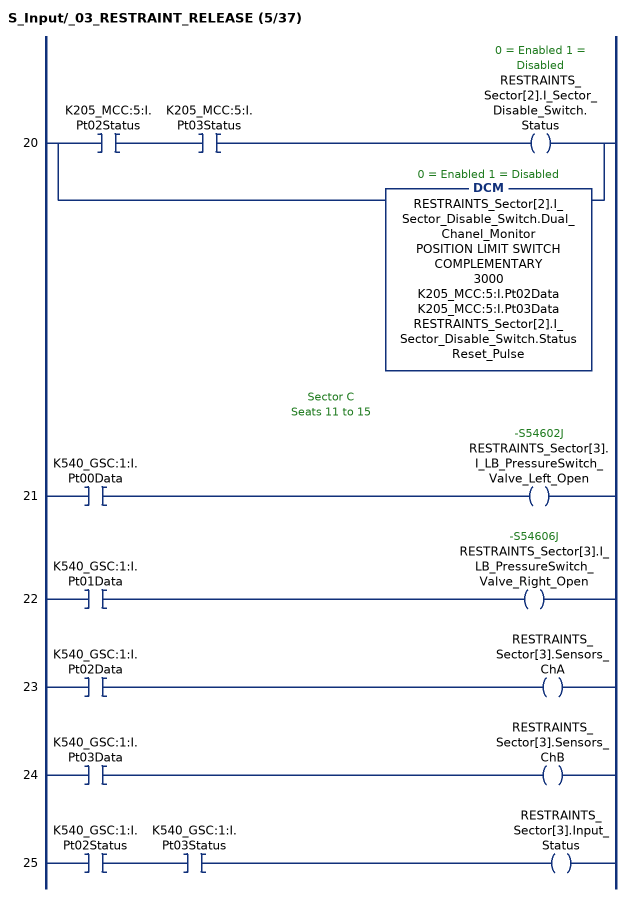
   20: [XIC(K205_MCC:5:I.Pt02Status) XIC(K205_MCC:5:I.Pt03Status) OTE(RESTRAINTS_Sector[2].I_Sector_Disable_Switch.Status) ,DCM(RESTRAINTS_Sector[2].I_Sector_Disable_Switch.Dual_Chanel_Monitor,POSITION LIMIT SWITCH,COMPLEMENTARY,3000,K205_MCC:5:I.Pt02Data,K205_MCC:5:I.Pt03Data,RESTRAINTS_Sector[2].I_Sector_Disable_Switch.Status,Reset_Pulse) ];
   // Sector C
   // Seats 11 to 15
   21: XIC(K540_GSC:1:I.Pt00Data)OTE(RESTRAINTS_Sector[3].I_LB_PressureSwitch_Valve_Left_Open);
   22: XIC(K540_GSC:1:I.Pt01Data)OTE(RESTRAINTS_Sector[3].I_LB_PressureSwitch_Valve_Right_Open);
   23: XIC(K540_GSC:1:I.Pt02Data)OTE(RESTRAINTS_Sector[3].Sensors_ChA);
   24: XIC(K540_GSC:1:I.Pt03Data)OTE(RESTRAINTS_Sector[3].Sensors_ChB);
   25: XIC(K540_GSC:1:I.Pt02Status)XIC(K540_GSC:1:I.Pt03Status)OTE(RESTRAINTS_Sector[3].Input_Status);
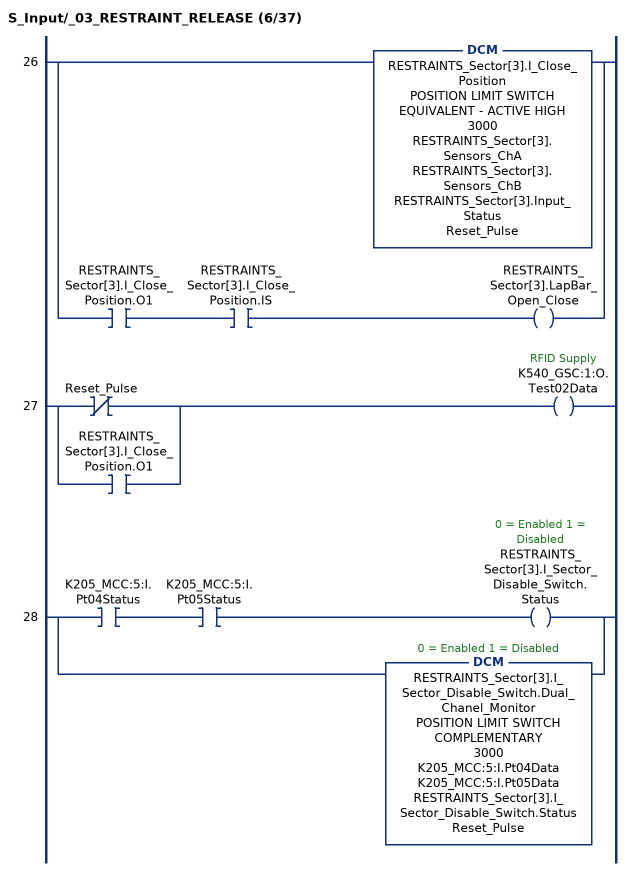
   26: [DCM(RESTRAINTS_Sector[3].I_Close_Position,POSITION LIMIT SWITCH,EQUIVALENT - ACTIVE HIGH,3000,RESTRAINTS_Sector[3].Sensors_ChA,RESTRAINTS_Sector[3].Sensors_ChB,RESTRAINTS_Sector[3].Input_Status,Reset_Pulse) ,XIC(RESTRAINTS_Sector[3].I_Close_Position.O1) XIC(RESTRAINTS_Sector[3].I_Close_Position.IS) OTE(RESTRAINTS_Sector[3].LapBar_Open_Close) ];
   27: [XIO(Reset_Pulse) ,XIC(RESTRAINTS_Sector[3].I_Close_Position.O1) ]OTE(K540_GSC:1:O.Test02Data);
   28: [XIC(K205_MCC:5:I.Pt04Status) XIC(K205_MCC:5:I.Pt05Status) OTE(RESTRAINTS_Sector[3].I_Sector_Disable_Switch.Status) ,DCM(RESTRAINTS_Sector[3].I_Sector_Disable_Switch.Dual_Chanel_Monitor,POSITION LIMIT SWITCH,COMPLEMENTARY,3000,K205_MCC:5:I.Pt04Data,K205_MCC:5:I.Pt05Data,RESTRAINTS_Sector[3].I_Sector_Disable_Switch.Status,Reset_Pulse) ];
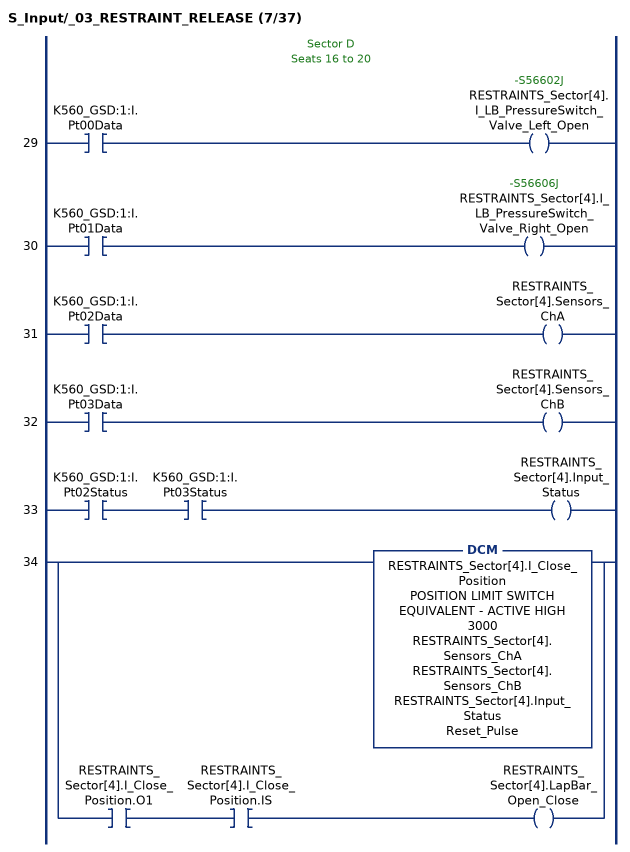
   // Sector D
   // Seats 16 to 20
   29: XIC(K560_GSD:1:I.Pt00Data)OTE(RESTRAINTS_Sector[4].I_LB_PressureSwitch_Valve_Left_Open);
   30: XIC(K560_GSD:1:I.Pt01Data)OTE(RESTRAINTS_Sector[4].I_LB_PressureSwitch_Valve_Right_Open);
   31: XIC(K560_GSD:1:I.Pt02Data)OTE(RESTRAINTS_Sector[4].Sensors_ChA);
   32: XIC(K560_GSD:1:I.Pt03Data)OTE(RESTRAINTS_Sector[4].Sensors_ChB);
   33: XIC(K560_GSD:1:I.Pt02Status)XIC(K560_GSD:1:I.Pt03Status)OTE(RESTRAINTS_Sector[4].Input_Status);
   34: [DCM(RESTRAINTS_Sector[4].I_Close_Position,POSITION LIMIT SWITCH,EQUIVALENT - ACTIVE HIGH,3000,RESTRAINTS_Sector[4].Sensors_ChA,RESTRAINTS_Sector[4].Sensors_ChB,RESTRAINTS_Sector[4].Input_Status,Reset_Pulse) ,XIC(RESTRAINTS_Sector[4].I_Close_Position.O1) XIC(RESTRAINTS_Sector[4].I_Close_Position.IS) OTE(RESTRAINTS_Sector[4].LapBar_Open_Close) ];
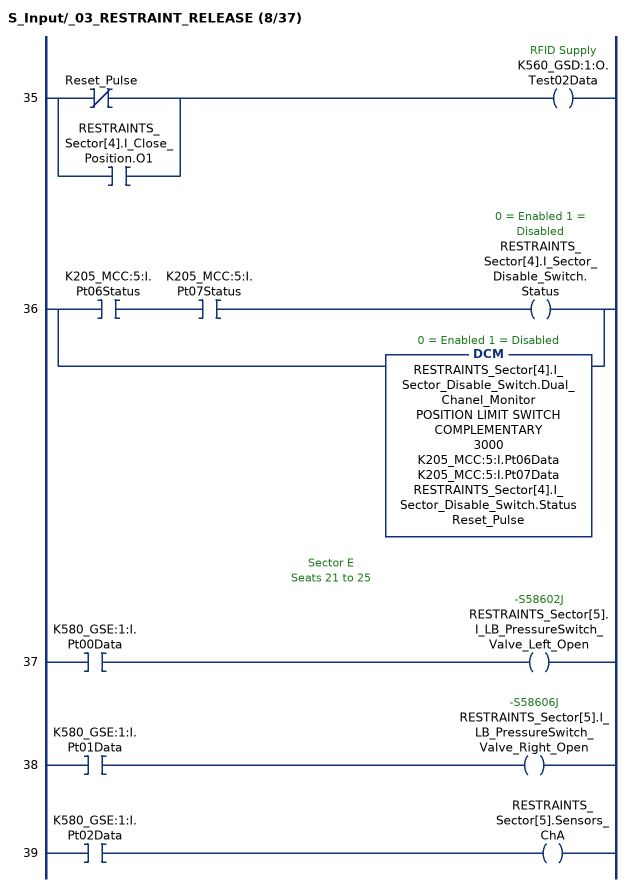
   35: [XIO(Reset_Pulse) ,XIC(RESTRAINTS_Sector[4].I_Close_Position.O1) ]OTE(K560_GSD:1:O.Test02Data);
   36: [XIC(K205_MCC:5:I.Pt06Status) XIC(K205_MCC:5:I.Pt07Status) OTE(RESTRAINTS_Sector[4].I_Sector_Disable_Switch.Status) ,DCM(RESTRAINTS_Sector[4].I_Sector_Disable_Switch.Dual_Chanel_Monitor,POSITION LIMIT SWITCH,COMPLEMENTARY,3000,K205_MCC:5:I.Pt06Data,K205_MCC:5:I.Pt07Data,RESTRAINTS_Sector[4].I_Sector_Disable_Switch.Status,Reset_Pulse) ];
   // Sector E
   // Seats 21 to 25
   37: XIC(K580_GSE:1:I.Pt00Data)OTE(RESTRAINTS_Sector[5].I_LB_PressureSwitch_Valve_Left_Open);
   38: XIC(K580_GSE:1:I.Pt01Data)OTE(RESTRAINTS_Sector[5].I_LB_PressureSwitch_Valve_Right_Open);
   39: XIC(K580_GSE:1:I.Pt02Data)OTE(RESTRAINTS_Sector[5].Sensors_ChA);
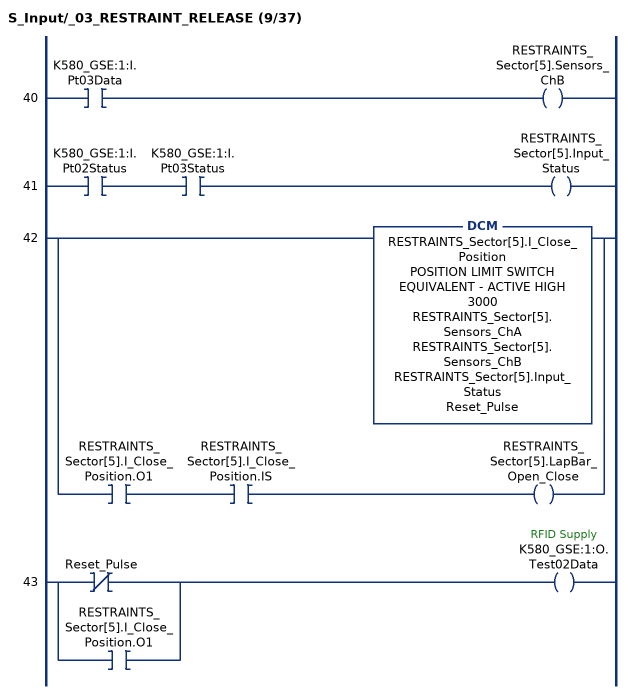
   40: XIC(K580_GSE:1:I.Pt03Data)OTE(RESTRAINTS_Sector[5].Sensors_ChB);
   41: XIC(K580_GSE:1:I.Pt02Status)XIC(K580_GSE:1:I.Pt03Status)OTE(RESTRAINTS_Sector[5].Input_Status);
   42: [DCM(RESTRAINTS_Sector[5].I_Close_Position,POSITION LIMIT SWITCH,EQUIVALENT - ACTIVE HIGH,3000,RESTRAINTS_Sector[5].Sensors_ChA,RESTRAINTS_Sector[5].Sensors_ChB,RESTRAINTS_Sector[5].Input_Status,Reset_Pulse) ,XIC(RESTRAINTS_Sector[5].I_Close_Position.O1) XIC(RESTRAINTS_Sector[5].I_Close_Position.IS) OTE(RESTRAINTS_Sector[5].LapBar_Open_Close) ];
   43: [XIO(Reset_Pulse) ,XIC(RESTRAINTS_Sector[5].I_Close_Position.O1) ]OTE(K580_GSE:1:O.Test02Data);
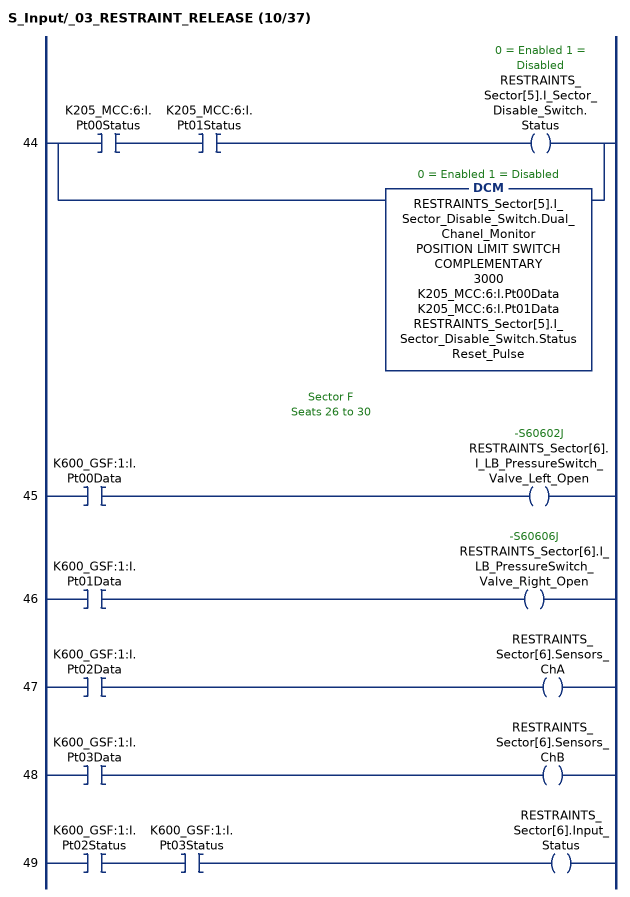
   44: [XIC(K205_MCC:6:I.Pt00Status) XIC(K205_MCC:6:I.Pt01Status) OTE(RESTRAINTS_Sector[5].I_Sector_Disable_Switch.Status) ,DCM(RESTRAINTS_Sector[5].I_Sector_Disable_Switch.Dual_Chanel_Monitor,POSITION LIMIT SWITCH,COMPLEMENTARY,3000,K205_MCC:6:I.Pt00Data,K205_MCC:6:I.Pt01Data,RESTRAINTS_Sector[5].I_Sector_Disable_Switch.Status,Reset_Pulse) ];
   // Sector F
   // Seats 26 to 30
   45: XIC(K600_GSF:1:I.Pt00Data)OTE(RESTRAINTS_Sector[6].I_LB_PressureSwitch_Valve_Left_Open);
   46: XIC(K600_GSF:1:I.Pt01Data)OTE(RESTRAINTS_Sector[6].I_LB_PressureSwitch_Valve_Right_Open);
   47: XIC(K600_GSF:1:I.Pt02Data)OTE(RESTRAINTS_Sector[6].Sensors_ChA);
   48: XIC(K600_GSF:1:I.Pt03Data)OTE(RESTRAINTS_Sector[6].Sensors_ChB);
   49: XIC(K600_GSF:1:I.Pt02Status)XIC(K600_GSF:1:I.Pt03Status)OTE(RESTRAINTS_Sector[6].Input_Status);
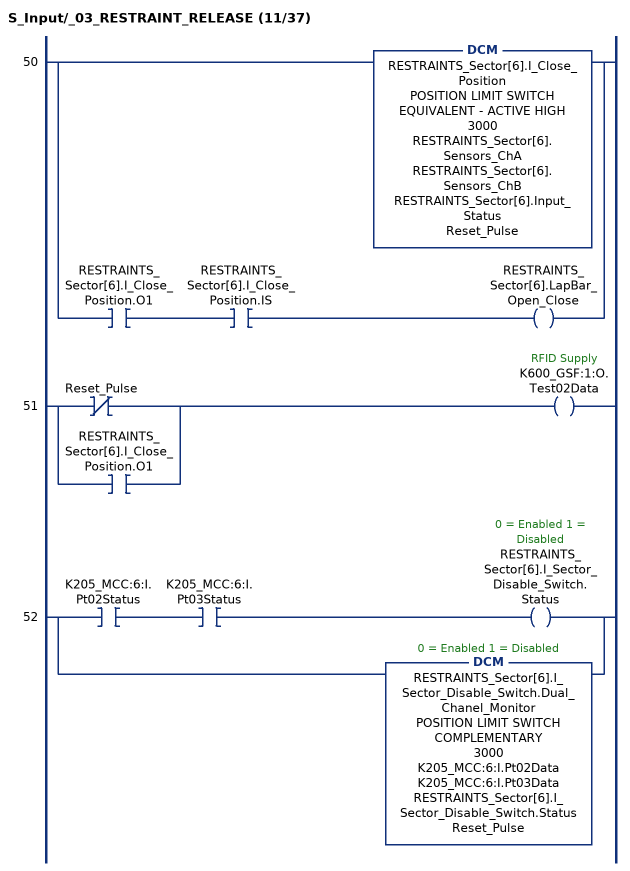
   50: [DCM(RESTRAINTS_Sector[6].I_Close_Position,POSITION LIMIT SWITCH,EQUIVALENT - ACTIVE HIGH,3000,RESTRAINTS_Sector[6].Sensors_ChA,RESTRAINTS_Sector[6].Sensors_ChB,RESTRAINTS_Sector[6].Input_Status,Reset_Pulse) ,XIC(RESTRAINTS_Sector[6].I_Close_Position.O1) XIC(RESTRAINTS_Sector[6].I_Close_Position.IS) OTE(RESTRAINTS_Sector[6].LapBar_Open_Close) ];
   51: [XIO(Reset_Pulse) ,XIC(RESTRAINTS_Sector[6].I_Close_Position.O1) ]OTE(K600_GSF:1:O.Test02Data);
   52: [XIC(K205_MCC:6:I.Pt02Status) XIC(K205_MCC:6:I.Pt03Status) OTE(RESTRAINTS_Sector[6].I_Sector_Disable_Switch.Status) ,DCM(RESTRAINTS_Sector[6].I_Sector_Disable_Switch.Dual_Chanel_Monitor,POSITION LIMIT SWITCH,COMPLEMENTARY,3000,K205_MCC:6:I.Pt02Data,K205_MCC:6:I.Pt03Data,RESTRAINTS_Sector[6].I_Sector_Disable_Switch.Status,Reset_Pulse) ];
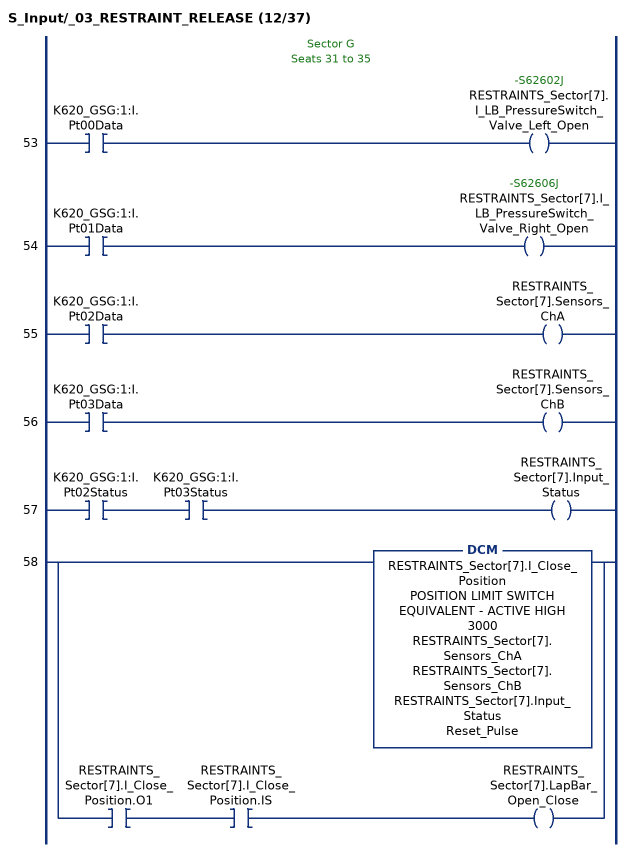
   // Sector G
   // Seats 31 to 35
   53: XIC(K620_GSG:1:I.Pt00Data)OTE(RESTRAINTS_Sector[7].I_LB_PressureSwitch_Valve_Left_Open);
   54: XIC(K620_GSG:1:I.Pt01Data)OTE(RESTRAINTS_Sector[7].I_LB_PressureSwitch_Valve_Right_Open);
   55: XIC(K620_GSG:1:I.Pt02Data)OTE(RESTRAINTS_Sector[7].Sensors_ChA);
   56: XIC(K620_GSG:1:I.Pt03Data)OTE(RESTRAINTS_Sector[7].Sensors_ChB);
   57: XIC(K620_GSG:1:I.Pt02Status)XIC(K620_GSG:1:I.Pt03Status)OTE(RESTRAINTS_Sector[7].Input_Status);
   58: [DCM(RESTRAINTS_Sector[7].I_Close_Position,POSITION LIMIT SWITCH,EQUIVALENT - ACTIVE HIGH,3000,RESTRAINTS_Sector[7].Sensors_ChA,RESTRAINTS_Sector[7].Sensors_ChB,RESTRAINTS_Sector[7].Input_Status,Reset_Pulse) ,XIC(RESTRAINTS_Sector[7].I_Close_Position.O1) XIC(RESTRAINTS_Sector[7].I_Close_Position.IS) OTE(RESTRAINTS_Sector[7].LapBar_Open_Close) ];
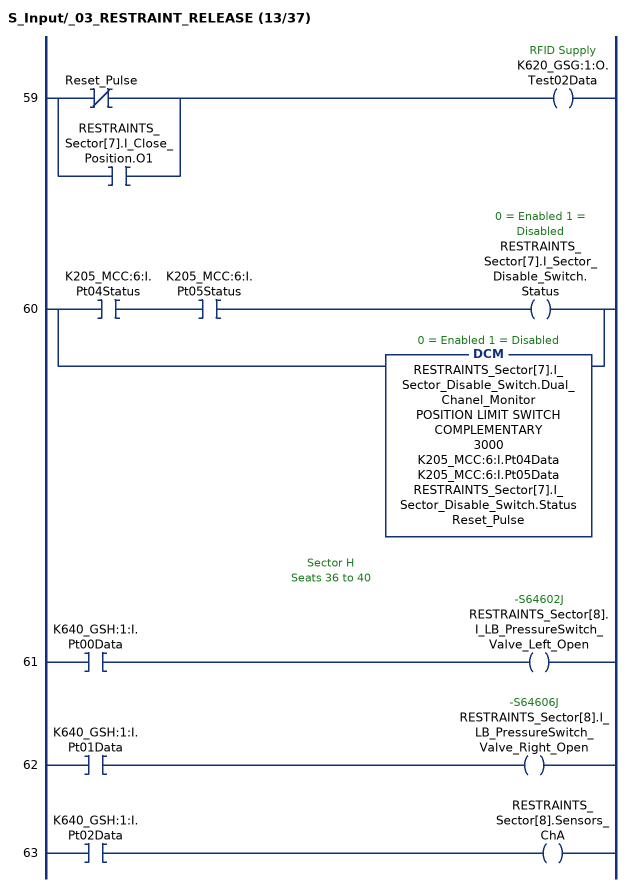
   59: [XIO(Reset_Pulse) ,XIC(RESTRAINTS_Sector[7].I_Close_Position.O1) ]OTE(K620_GSG:1:O.Test02Data);
   60: [XIC(K205_MCC:6:I.Pt04Status) XIC(K205_MCC:6:I.Pt05Status) OTE(RESTRAINTS_Sector[7].I_Sector_Disable_Switch.Status) ,DCM(RESTRAINTS_Sector[7].I_Sector_Disable_Switch.Dual_Chanel_Monitor,POSITION LIMIT SWITCH,COMPLEMENTARY,3000,K205_MCC:6:I.Pt04Data,K205_MCC:6:I.Pt05Data,RESTRAINTS_Sector[7].I_Sector_Disable_Switch.Status,Reset_Pulse) ];
   // Sector H
   // Seats 36 to 40
   61: XIC(K640_GSH:1:I.Pt00Data)OTE(RESTRAINTS_Sector[8].I_LB_PressureSwitch_Valve_Left_Open);
   62: XIC(K640_GSH:1:I.Pt01Data)OTE(RESTRAINTS_Sector[8].I_LB_PressureSwitch_Valve_Right_Open);
   63: XIC(K640_GSH:1:I.Pt02Data)OTE(RESTRAINTS_Sector[8].Sensors_ChA);
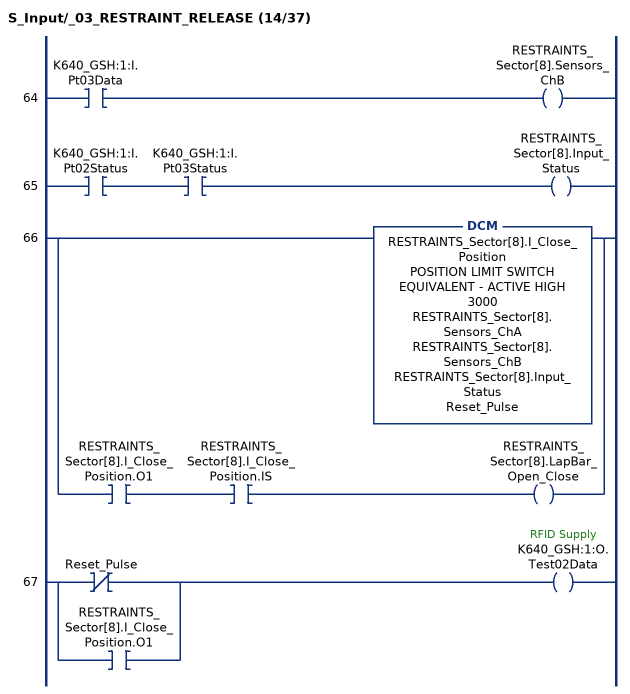
   64: XIC(K640_GSH:1:I.Pt03Data)OTE(RESTRAINTS_Sector[8].Sensors_ChB);
   65: XIC(K640_GSH:1:I.Pt02Status)XIC(K640_GSH:1:I.Pt03Status)OTE(RESTRAINTS_Sector[8].Input_Status);
   66: [DCM(RESTRAINTS_Sector[8].I_Close_Position,POSITION LIMIT SWITCH,EQUIVALENT - ACTIVE HIGH,3000,RESTRAINTS_Sector[8].Sensors_ChA,RESTRAINTS_Sector[8].Sensors_ChB,RESTRAINTS_Sector[8].Input_Status,Reset_Pulse) ,XIC(RESTRAINTS_Sector[8].I_Close_Position.O1) XIC(RESTRAINTS_Sector[8].I_Close_Position.IS) OTE(RESTRAINTS_Sector[8].LapBar_Open_Close) ];
   67: [XIO(Reset_Pulse) ,XIC(RESTRAINTS_Sector[8].I_Close_Position.O1) ]OTE(K640_GSH:1:O.Test02Data);
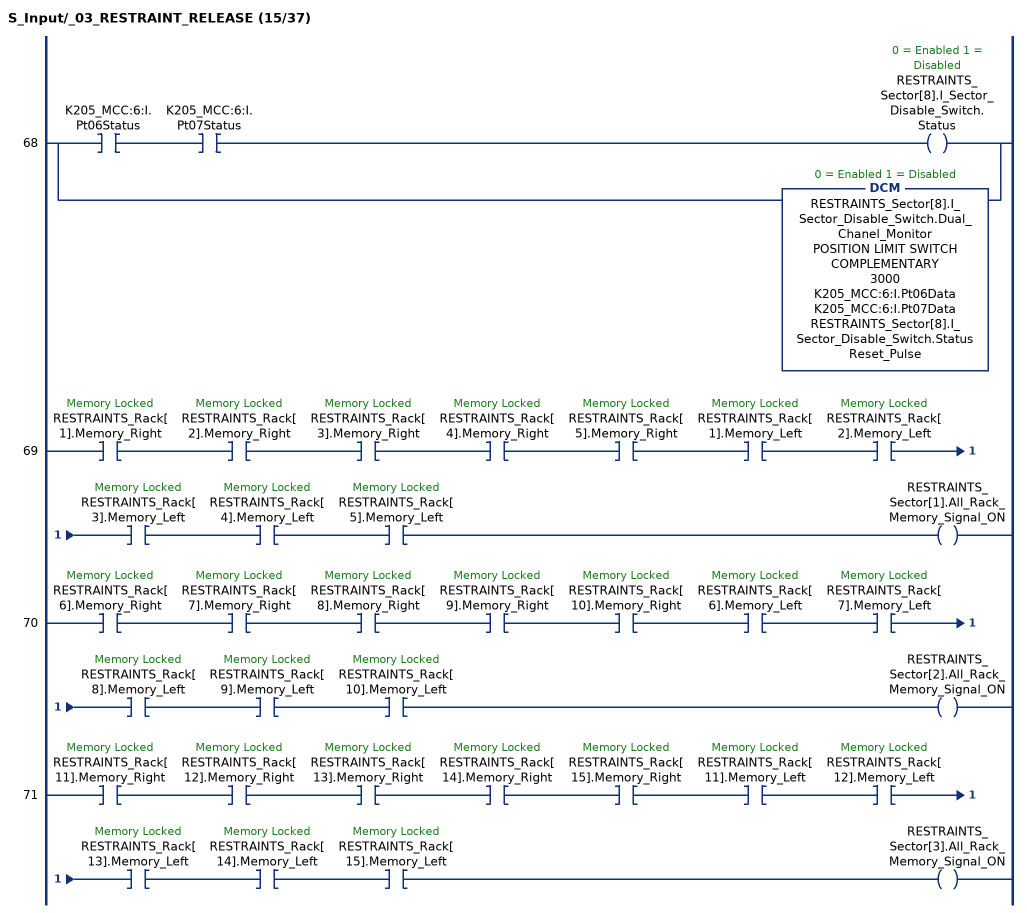
   68: [XIC(K205_MCC:6:I.Pt06Status) XIC(K205_MCC:6:I.Pt07Status) OTE(RESTRAINTS_Sector[8].I_Sector_Disable_Switch.Status) ,DCM(RESTRAINTS_Sector[8].I_Sector_Disable_Switch.Dual_Chanel_Monitor,POSITION LIMIT SWITCH,COMPLEMENTARY,3000,K205_MCC:6:I.Pt06Data,K205_MCC:6:I.Pt07Data,RESTRAINTS_Sector[8].I_Sector_Disable_Switch.Status,Reset_Pulse) ];
   69: XIC(RESTRAINTS_Rack[1].Memory_Right)XIC(RESTRAINTS_Rack[2].Memory_Right)XIC(RESTRAINTS_Rack[3].Memory_Right)XIC(RESTRAINTS_Rack[4].Memory_Right)XIC(RESTRAINTS_Rack[5].Memory_Right)XIC(RESTRAINTS_Rack[1].Memory_Left)XIC(RESTRAINTS_Rack[2].Memory_Left)XIC(RESTRAINTS_Rack[3].Memory_Left)XIC(RESTRAINTS_Rack[4].Memory_Left)XIC(RESTRAINTS_Rack[5].Memory_Left)OTE(RESTRAINTS_Sector[1].All_Rack_Memory_Signal_ON);
   70: XIC(RESTRAINTS_Rack[6].Memory_Right)XIC(RESTRAINTS_Rack[7].Memory_Right)XIC(RESTRAINTS_Rack[8].Memory_Right)XIC(RESTRAINTS_Rack[9].Memory_Right)XIC(RESTRAINTS_Rack[10].Memory_Right)XIC(RESTRAINTS_Rack[6].Memory_Left)XIC(RESTRAINTS_Rack[7].Memory_Left)XIC(RESTRAINTS_Rack[8].Memory_Left)XIC(RESTRAINTS_Rack[9].Memory_Left)XIC(RESTRAINTS_Rack[10].Memory_Left)OTE(RESTRAINTS_Sector[2].All_Rack_Memory_Signal_ON);
   71: XIC(RESTRAINTS_Rack[11].Memory_Right)XIC(RESTRAINTS_Rack[12].Memory_Right)XIC(RESTRAINTS_Rack[13].Memory_Right)XIC(RESTRAINTS_Rack[14].Memory_Right)XIC(RESTRAINTS_Rack[15].Memory_Right)XIC(RESTRAINTS_Rack[11].Memory_Left)XIC(RESTRAINTS_Rack[12].Memory_Left)XIC(RESTRAINTS_Rack[13].Memory_Left)XIC(RESTRAINTS_Rack[14].Memory_Left)XIC(RESTRAINTS_Rack[15].Memory_Left)OTE(RESTRAINTS_Sector[3].All_Rack_Memory_Signal_ON);
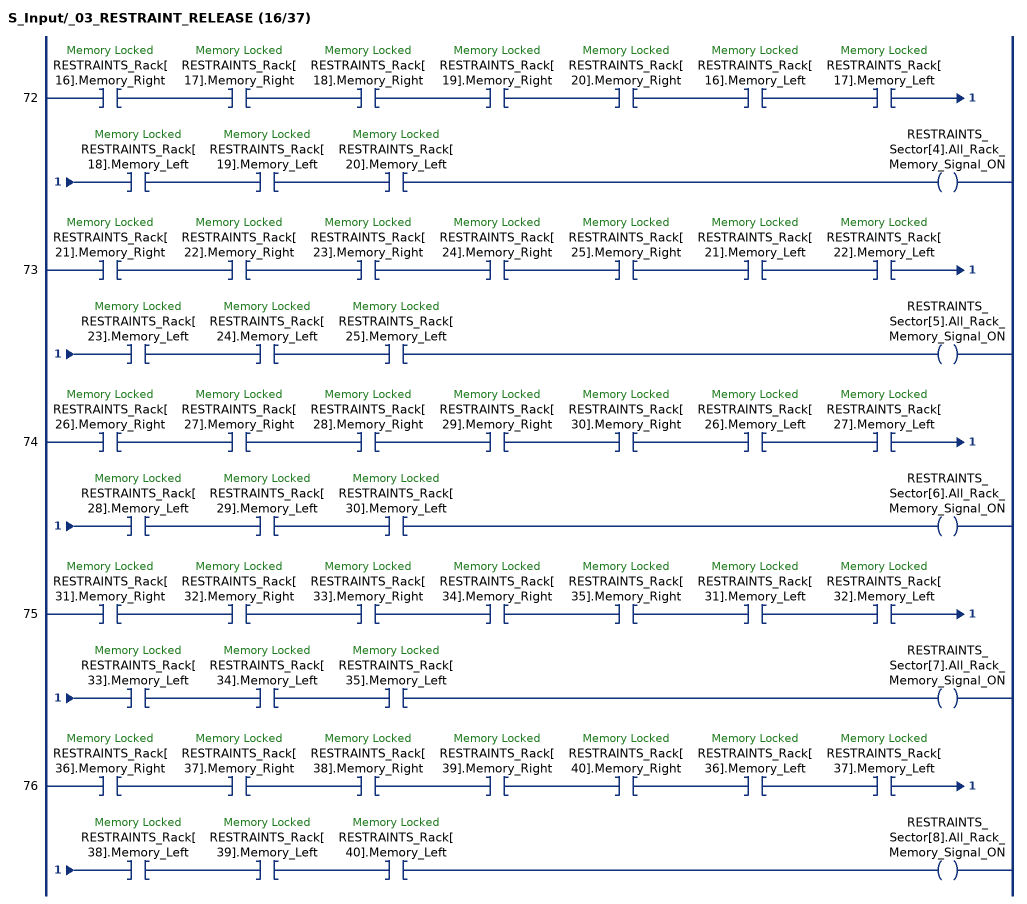
   72: XIC(RESTRAINTS_Rack[16].Memory_Right)XIC(RESTRAINTS_Rack[17].Memory_Right)XIC(RESTRAINTS_Rack[18].Memory_Right)XIC(RESTRAINTS_Rack[19].Memory_Right)XIC(RESTRAINTS_Rack[20].Memory_Right)XIC(RESTRAINTS_Rack[16].Memory_Left)XIC(RESTRAINTS_Rack[17].Memory_Left)XIC(RESTRAINTS_Rack[18].Memory_Left)XIC(RESTRAINTS_Rack[19].Memory_Left)XIC(RESTRAINTS_Rack[20].Memory_Left)OTE(RESTRAINTS_Sector[4].All_Rack_Memory_Signal_ON);
   73: XIC(RESTRAINTS_Rack[21].Memory_Right)XIC(RESTRAINTS_Rack[22].Memory_Right)XIC(RESTRAINTS_Rack[23].Memory_Right)XIC(RESTRAINTS_Rack[24].Memory_Right)XIC(RESTRAINTS_Rack[25].Memory_Right)XIC(RESTRAINTS_Rack[21].Memory_Left)XIC(RESTRAINTS_Rack[22].Memory_Left)XIC(RESTRAINTS_Rack[23].Memory_Left)XIC(RESTRAINTS_Rack[24].Memory_Left)XIC(RESTRAINTS_Rack[25].Memory_Left)OTE(RESTRAINTS_Sector[5].All_Rack_Memory_Signal_ON);
   74: XIC(RESTRAINTS_Rack[26].Memory_Right)XIC(RESTRAINTS_Rack[27].Memory_Right)XIC(RESTRAINTS_Rack[28].Memory_Right)XIC(RESTRAINTS_Rack[29].Memory_Right)XIC(RESTRAINTS_Rack[30].Memory_Right)XIC(RESTRAINTS_Rack[26].Memory_Left)XIC(RESTRAINTS_Rack[27].Memory_Left)XIC(RESTRAINTS_Rack[28].Memory_Left)XIC(RESTRAINTS_Rack[29].Memory_Left)XIC(RESTRAINTS_Rack[30].Memory_Left)OTE(RESTRAINTS_Sector[6].All_Rack_Memory_Signal_ON);
   75: XIC(RESTRAINTS_Rack[31].Memory_Right)XIC(RESTRAINTS_Rack[32].Memory_Right)XIC(RESTRAINTS_Rack[33].Memory_Right)XIC(RESTRAINTS_Rack[34].Memory_Right)XIC(RESTRAINTS_Rack[35].Memory_Right)XIC(RESTRAINTS_Rack[31].Memory_Left)XIC(RESTRAINTS_Rack[32].Memory_Left)XIC(RESTRAINTS_Rack[33].Memory_Left)XIC(RESTRAINTS_Rack[34].Memory_Left)XIC(RESTRAINTS_Rack[35].Memory_Left)OTE(RESTRAINTS_Sector[7].All_Rack_Memory_Signal_ON);
   76: XIC(RESTRAINTS_Rack[36].Memory_Right)XIC(RESTRAINTS_Rack[37].Memory_Right)XIC(RESTRAINTS_Rack[38].Memory_Right)XIC(RESTRAINTS_Rack[39].Memory_Right)XIC(RESTRAINTS_Rack[40].Memory_Right)XIC(RESTRAINTS_Rack[36].Memory_Left)XIC(RESTRAINTS_Rack[37].Memory_Left)XIC(RESTRAINTS_Rack[38].Memory_Left)XIC(RESTRAINTS_Rack[39].Memory_Left)XIC(RESTRAINTS_Rack[40].Memory_Left)OTE(RESTRAINTS_Sector[8].All_Rack_Memory_Signal_ON);
